(* Logix 5000 project; controller PLC_MCC1300_75F1 vendor 1 type 14 code 166 rev 32.11; software revision 32.04; part 83 of 83 *)
(* tags used below, declared in another part *)
   GP_OB_InitializeMain : GP_OB_Initialize;
   M302SpeedUp : MAC_SpeedUp;
   M360_M1_DR : AXIS_CIP_DRIVE;
   TMP_dDirection : DINT;
   TMP_dTarget : DINT;
   TMP_rAcc : REAL;
   TMP_rDec : REAL;
   TMP_rSpeed : REAL;
   Z300_Conveyor : UDT_StandConv[29];
   Z300_Conveyor_IN_MOTION : MAC_Conveyor_ZC_IN_MOTION[29];
   Z300_Conveyor_OUT_MOTION : MAC_Conveyor_ZC_OUT_MOTION[29];
(* MotionLogic, continued *)

ROUTINE M360_Motion   (* ladder *)
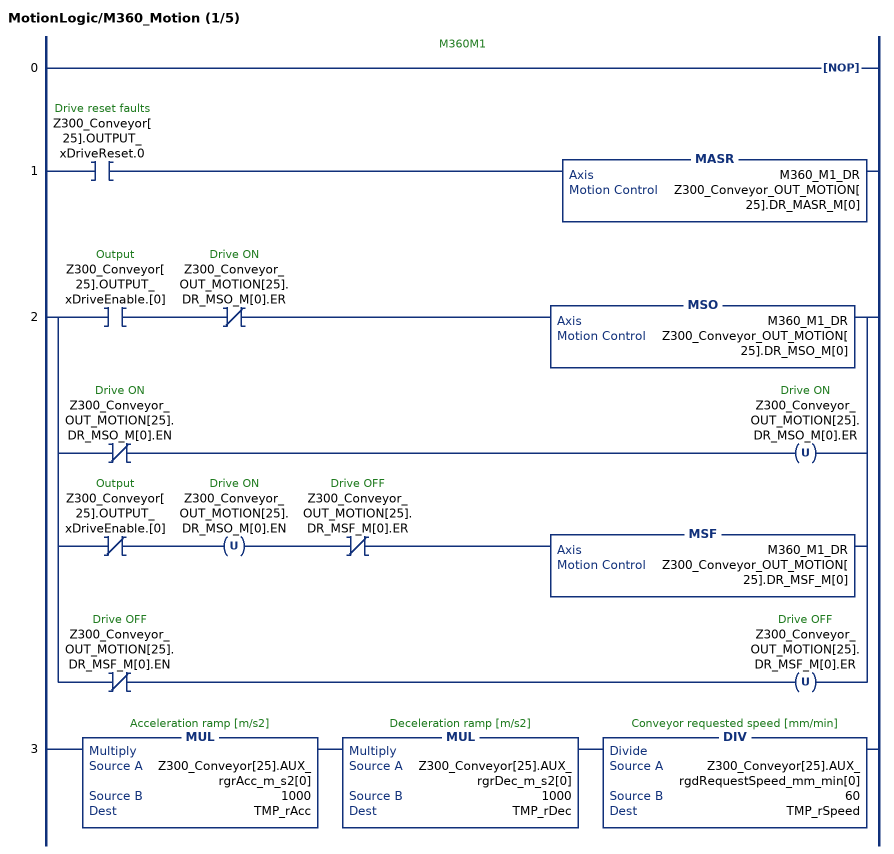
   // M360M1
   0: NOP();
   1: XIC(Z300_Conveyor[25].OUTPUT_xDriveReset.0)MASR(M360_M1_DR,Z300_Conveyor_OUT_MOTION[25].DR_MASR_M[0]);
   2: [XIC(Z300_Conveyor[25].OUTPUT_xDriveEnable.[0]) XIO(Z300_Conveyor_OUT_MOTION[25].DR_MSO_M[0].ER) MSO(M360_M1_DR,Z300_Conveyor_OUT_MOTION[25].DR_MSO_M[0]) ,XIO(Z300_Conveyor_OUT_MOTION[25].DR_MSO_M[0].EN) OTU(Z300_Conveyor_OUT_MOTION[25].DR_MSO_M[0].ER) ,XIO(Z300_Conveyor[25].OUTPUT_xDriveEnable.[0]) OTU(Z300_Conveyor_OUT_MOTION[25].DR_MSO_M[0].EN) XIO(Z300_Conveyor_OUT_MOTION[25].DR_MSF_M[0].ER) MSF(M360_M1_DR,Z300_Conveyor_OUT_MOTION[25].DR_MSF_M[0]) ,XIO(Z300_Conveyor_OUT_MOTION[25].DR_MSF_M[0].EN) OTU(Z300_Conveyor_OUT_MOTION[25].DR_MSF_M[0].ER) ];
   3: MUL(Z300_Conveyor[25].AUX_rgrAcc_m_s2[0],1000,TMP_rAcc)MUL(Z300_Conveyor[25].AUX_rgrDec_m_s2[0],1000,TMP_rDec)DIV(Z300_Conveyor[25].AUX_rgdRequestSpeed_mm_min[0],60,TMP_rSpeed);
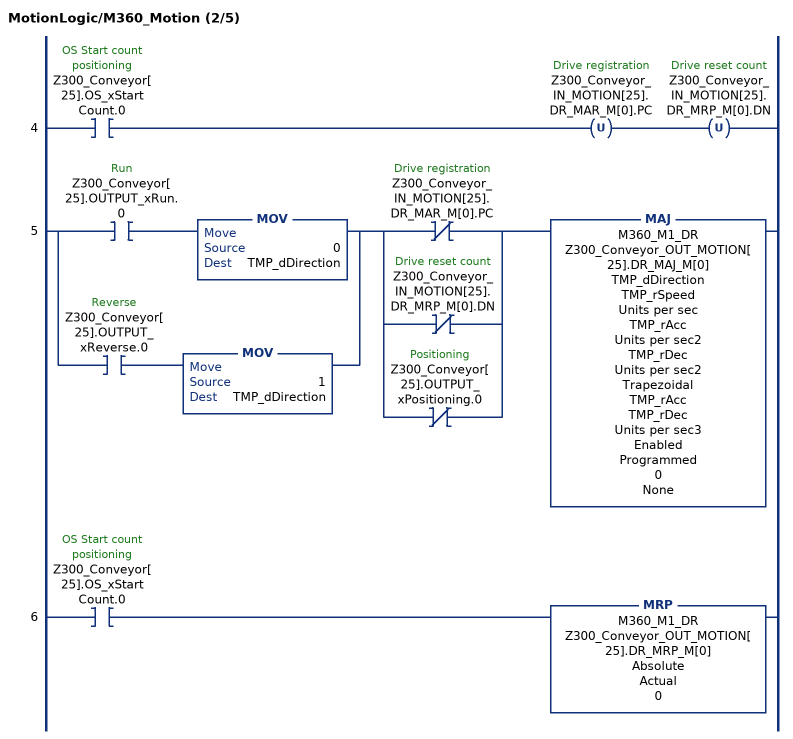
   4: XIC(Z300_Conveyor[25].OS_xStartCount.0)OTU(Z300_Conveyor_IN_MOTION[25].DR_MAR_M[0].PC)OTU(Z300_Conveyor_IN_MOTION[25].DR_MRP_M[0].DN);
   5: [XIC(Z300_Conveyor[25].OUTPUT_xRun.0) MOV(0,TMP_dDirection) ,XIC(Z300_Conveyor[25].OUTPUT_xReverse.0) MOV(1,TMP_dDirection) ][XIO(Z300_Conveyor_IN_MOTION[25].DR_MAR_M[0].PC) ,XIO(Z300_Conveyor_IN_MOTION[25].DR_MRP_M[0].DN) ,XIO(Z300_Conveyor[25].OUTPUT_xPositioning.0) ]MAJ(M360_M1_DR,Z300_Conveyor_OUT_MOTION[25].DR_MAJ_M[0],TMP_dDirection,TMP_rSpeed,Units per sec,TMP_rAcc,Units per sec2,TMP_rDec,Units per sec2,Trapezoidal,TMP_rAcc,TMP_rDec,Units per sec3,Enabled,Programmed,0,None);
   6: XIC(Z300_Conveyor[25].OS_xStartCount.0)MRP(M360_M1_DR,Z300_Conveyor_OUT_MOTION[25].DR_MRP_M[0],Absolute,Actual,0);
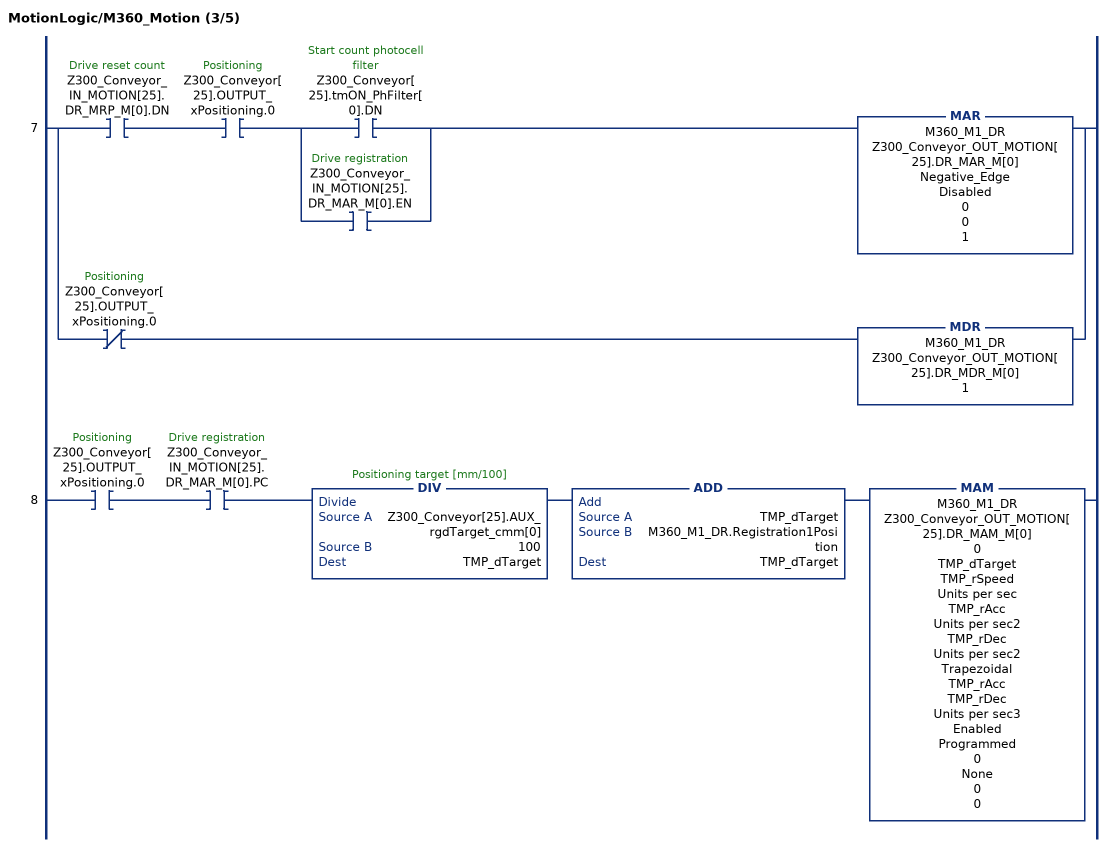
   7: [XIC(Z300_Conveyor_IN_MOTION[25].DR_MRP_M[0].DN) XIC(Z300_Conveyor[25].OUTPUT_xPositioning.0) [XIC(Z300_Conveyor[25].tmON_PhFilter[0].DN) ,XIC(Z300_Conveyor_IN_MOTION[25].DR_MAR_M[0].EN) ] MAR(M360_M1_DR,Z300_Conveyor_OUT_MOTION[25].DR_MAR_M[0],Negative_Edge,Disabled,0,0,1) ,XIO(Z300_Conveyor[25].OUTPUT_xPositioning.0) MDR(M360_M1_DR,Z300_Conveyor_OUT_MOTION[25].DR_MDR_M[0],1) ];
   8: XIC(Z300_Conveyor[25].OUTPUT_xPositioning.0)XIC(Z300_Conveyor_IN_MOTION[25].DR_MAR_M[0].PC)DIV(Z300_Conveyor[25].AUX_rgdTarget_cmm[0],100,TMP_dTarget)ADD(TMP_dTarget,M360_M1_DR.Registration1Position,TMP_dTarget)MAM(M360_M1_DR,Z300_Conveyor_OUT_MOTION[25].DR_MAM_M[0],0,TMP_dTarget,TMP_rSpeed,Units per sec,TMP_rAcc,Units per sec2,TMP_rDec,Units per sec2,Trapezoidal,TMP_rAcc,TMP_rDec,Units per sec3,Enabled,Programmed,0,None,0,0);
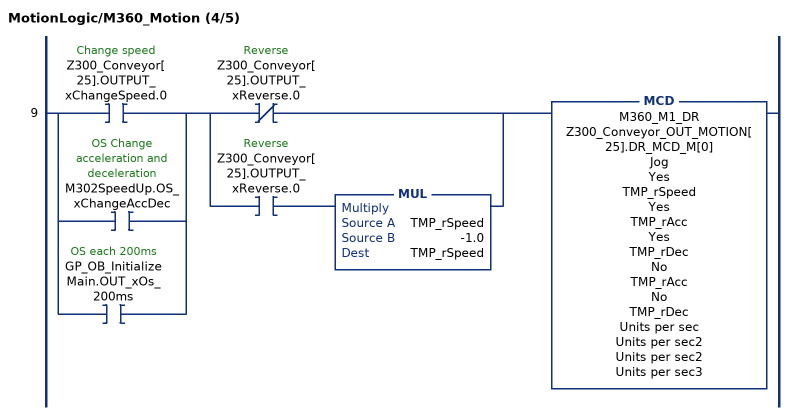
   9: [XIC(Z300_Conveyor[25].OUTPUT_xChangeSpeed.0) ,XIC(M302SpeedUp.OS_xChangeAccDec) ,XIC(GP_OB_InitializeMain.OUT_xOs_200ms) ][XIO(Z300_Conveyor[25].OUTPUT_xReverse.0) ,XIC(Z300_Conveyor[25].OUTPUT_xReverse.0) MUL(TMP_rSpeed,-1.0,TMP_rSpeed) ]MCD(M360_M1_DR,Z300_Conveyor_OUT_MOTION[25].DR_MCD_M[0],Jog,Yes,TMP_rSpeed,Yes,TMP_rAcc,Yes,TMP_rDec,No,TMP_rAcc,No,TMP_rDec,Units per sec,Units per sec2,Units per sec2,Units per sec3);
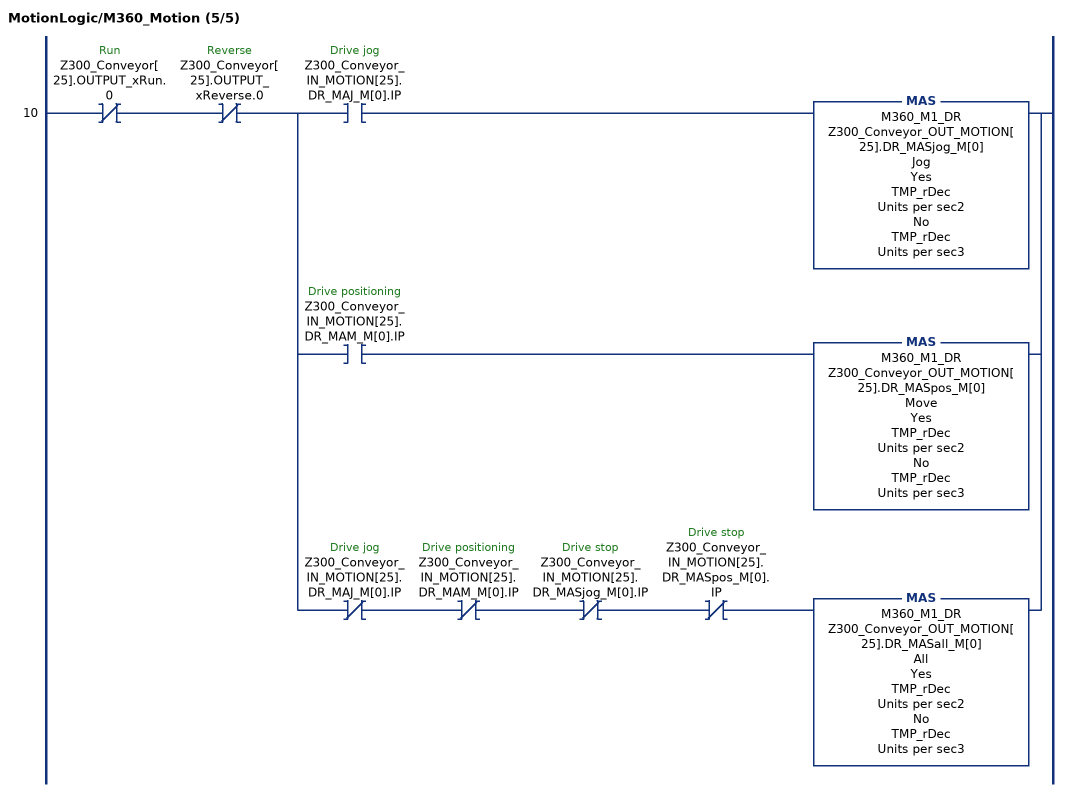
   10: XIO(Z300_Conveyor[25].OUTPUT_xRun.0)XIO(Z300_Conveyor[25].OUTPUT_xReverse.0)[XIC(Z300_Conveyor_IN_MOTION[25].DR_MAJ_M[0].IP) MAS(M360_M1_DR,Z300_Conveyor_OUT_MOTION[25].DR_MASjog_M[0],Jog,Yes,TMP_rDec,Units per sec2,No,TMP_rDec,Units per sec3) ,XIC(Z300_Conveyor_IN_MOTION[25].DR_MAM_M[0].IP) MAS(M360_M1_DR,Z300_Conveyor_OUT_MOTION[25].DR_MASpos_M[0],Move,Yes,TMP_rDec,Units per sec2,No,TMP_rDec,Units per sec3) ,XIO(Z300_Conveyor_IN_MOTION[25].DR_MAJ_M[0].IP) XIO(Z300_Conveyor_IN_MOTION[25].DR_MAM_M[0].IP) XIO(Z300_Conveyor_IN_MOTION[25].DR_MASjog_M[0].IP) XIO(Z300_Conveyor_IN_MOTION[25].DR_MASpos_M[0].IP) MAS(M360_M1_DR,Z300_Conveyor_OUT_MOTION[25].DR_MASall_M[0],All,Yes,TMP_rDec,Units per sec2,No,TMP_rDec,Units per sec3) ];
END_ROUTINE

ROUTINE Main   (* ladder *)
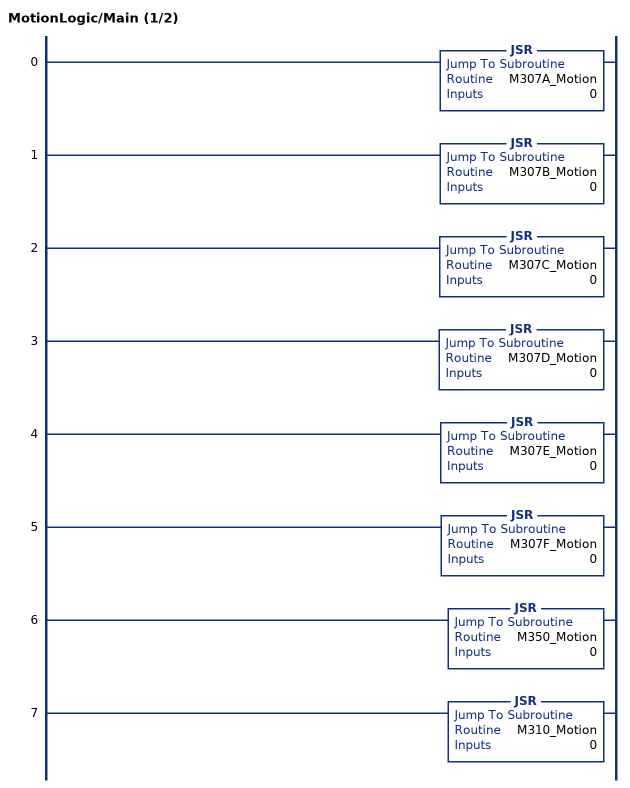
   0: JSR(M307A_Motion,0);
   1: JSR(M307B_Motion,0);
   2: JSR(M307C_Motion,0);
   3: JSR(M307D_Motion,0);
   4: JSR(M307E_Motion,0);
   5: JSR(M307F_Motion,0);
   6: JSR(M350_Motion,0);
   7: JSR(M310_Motion,0);
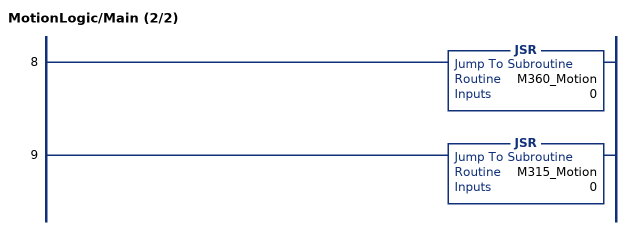
   8: JSR(M360_Motion,0);
   9: JSR(M315_Motion,0);
END_ROUTINE
END_PROGRAM
